REGION Network 8: Control the filling valve
         A     #Temp_IO_Status.HM_FillingValve;
         S     #Temp_IO_Status.HM_FillingValve1;
         S     #Temp_IO_Status.HM_FillingValve2;
   //
         AN    #Temp_IO_Status.HM_FillingValve;
         AN    #IN_Max_Level_Tank;
         R     #Temp_IO_Status.HM_FillingValve1;
         R     #Temp_IO_Status.HM_FillingValve2;
   //
         AN    #Temp_IO_Status.HM_FillingValve;
         AN    #Temp_IO_Status.HMFillingValves_Open;
         A     #Temp_IO_Status.V_FillingValve1;
         A     #Temp_IO_Status.V_FillingValve2;
         S     #Temp_IO_Status.HMFillingValves_Open;
   //
         A     #Temp_IO_Status.HMFillingValves_Open;
         L     S5T#3S;
         SP    #IN_Timer_Overlap_Valves;
   //
         AN    #Temp_IO_Status.HM_FillingValve;
         A     #Temp_IO_Status.V_FillingValve1;
         A     #Temp_IO_Status.V_FillingValve2;
         A     #Temp_IO_Status.HMFillingValves_Open;
         AN    #IN_Timer_Overlap_Valves;
         R     #Temp_IO_Status.HMFillingValves_Open;
   //
         AN    #Temp_IO_Status.HM_FillingValve;
         A     #Temp_IO_Status.HMFillingValves_Open;
         R     #Temp_IO_Status.HM_FillingValve1;
   //
         AN    #Temp_IO_Status.HM_FillingValve;
         AN    #Temp_IO_Status.HMFillingValves_Open;
         R     #Temp_IO_Status.HM_FillingValve2;
   //
         A     #Temp_IO_Status.HM_FillingValve1;
         L     S5T#2S;
         SF    #IN_Timer_Valve1;
   //
         A     #IN_Timer_Valve1;
         =     #Temp_IO_Status.V_FillingValve1;
   //
         A     #Temp_IO_Status.HM_FillingValve2;
         L     S5T#2S;
         SF    #IN_Timer_Valve2;
   //
         A     #IN_Timer_Valve2;
         =     #Temp_IO_Status.V_FillingValve2;
   //
         A     #Temp_IO_Status.V_FillingValve1;
         =     #OUT_FillingValve1;
   //
         A     #Temp_IO_Status.V_FillingValve2;
         =     #OUT_FillingValve2;
END_REGION

REGION Network 9
         AN    #Temp_IO_Status.V_FillingValve1;
   //    U     "E_FuellVent1_K1_geschl"
         AN    #Temp_IO_Status.HM_Valve2_closed;
         S     #Temp_IO_Status.HM_Valve1_closed;
   //
         AN    #Temp_IO_Status.V_FillingValve2;
   //    U     "E_FuellVent2_K1_geschl"
         AN    #Temp_IO_Status.HM_Valve1_closed;
         S     #Temp_IO_Status.HM_Valve2_closed;
   //
         A     #Temp_IO_Status.V_FillingValve1;
   //    U     "E_FuellVent1_K1_offen"
         R     #Temp_IO_Status.HM_Valve1_closed;
   //
         A     #Temp_IO_Status.V_FillingValve2;
   //    U     "E_FuellVent2_K1_offen"
         R     #Temp_IO_Status.HM_Valve1_closed;
   //
         A     #Temp_IO_Status.EnableComponentPump;
         AN    #IN_Max_Level_Tank;
         AN    #Temp_IO_Fault.FLT_Valve1_Max;
         S     #Temp_IO_Fault.FLT_Valve1_Max;
         S     #IO_FaultLevel_3;
   //-----
         A     #Temp_IO_Status.HM_Valve2_closed;
         AN    #IN_Max_Level_Tank;
         AN    #Temp_IO_Fault.FLT_Valve2_Max;
         S     #Temp_IO_Fault.FLT_Valve2_Max;
         S     #IO_FaultLevel_3;
   //-----
END_REGION

REGION Network 10: Save data
   Out:  NOP   0;
         CALL  BLKMOV
         ( SRCBLK  := #Temp_IO_Status,
           RET_VAL := #ERROR_CODE,
           DSTBLK  := #AnyPointer1
         );
   //-----
         CALL  BLKMOV
         ( SRCBLK  := #Temp_IO_Fault,
           RET_VAL := #ERROR_CODE,
           DSTBLK  := #AnyPointer2
         );
   //-----
END_REGION
END_FUNCTION

FUNCTION "Baustein_1" : Void   // FC3, SCL
{ S7_Optimized_Access := 'FALSE' }
VERSION : 0.1
   VAR_TEMP
      N : Int;
      Y : Int;
   END_VAR
BEGIN

   // Anzahl der Komponenten am Mischkopf und Zuweisung der Namen vom Tagesbehälter!
   // 
     "DB619_State_MPart".Recirculation[1].Lowpressure_Exist := 0;
     "DB619_State_MPart".Recirculation[2].Lowpressure_Exist := 0;

   FOR #N := 1 TO "DB790_PlantParameter".AmountMH DO
     // Statement section FOR

   "DB704_MH_Value".Mixinghead[#N].MH_Connection[1].Exist:=0;
   "DB704_MH_Value".Mixinghead[#N].MH_Connection[2].Exist:=0;
   "DB704_MH_Value".Mixinghead[#N].MH_Connection[3].Exist:=0;
   "DB704_MH_Value".Mixinghead[#N].MH_Connection[4].Exist:=0;
   "DB704_MH_Value".Mixinghead[#N].MH_Connection[5].Exist:=0;
   "DB704_MH_Value".Mixinghead[#N].MH_Connection[6].Exist:=0;

     IF "DB704_MH_Value".Mixinghead[#N].AmountComponent = 1 THEN
       "DB704_MH_Value".Mixinghead[#N].MH_Connection[1].Exist:=1;
     ELSIF "DB704_MH_Value".Mixinghead[#N].AmountComponent = 2 THEN
       "DB704_MH_Value".Mixinghead[#N].MH_Connection[1].Exist:=1; 
       "DB704_MH_Value".Mixinghead[#N].MH_Connection[2].Exist:=1;
     ELSIF "DB704_MH_Value".Mixinghead[#N].AmountComponent = 3 THEN
       "DB704_MH_Value".Mixinghead[#N].MH_Connection[1].Exist:=1;
       "DB704_MH_Value".Mixinghead[#N].MH_Connection[2].Exist:=1;
       "DB704_MH_Value".Mixinghead[#N].MH_Connection[3].Exist:=1;
     ELSIF "DB704_MH_Value".Mixinghead[#N].AmountComponent = 4 THEN
       "DB704_MH_Value".Mixinghead[#N].MH_Connection[1].Exist:=1; 
       "DB704_MH_Value".Mixinghead[#N].MH_Connection[2].Exist:=1;
       "DB704_MH_Value".Mixinghead[#N].MH_Connection[3].Exist:=1;
       "DB704_MH_Value".Mixinghead[#N].MH_Connection[4].Exist:=1;
     ELSIF "DB704_MH_Value".Mixinghead[#N].AmountComponent = 5 THEN
       "DB704_MH_Value".Mixinghead[#N].MH_Connection[1].Exist:=1;
       "DB704_MH_Value".Mixinghead[#N].MH_Connection[2].Exist:=1;
       "DB704_MH_Value".Mixinghead[#N].MH_Connection[3].Exist:=1;
       "DB704_MH_Value".Mixinghead[#N].MH_Connection[4].Exist:=1;
       "DB704_MH_Value".Mixinghead[#N].MH_Connection[5].Exist:=1;
     ELSIF "DB704_MH_Value".Mixinghead[#N].AmountComponent = 6 THEN
       "DB704_MH_Value".Mixinghead[#N].MH_Connection[1].Exist:=1;
       "DB704_MH_Value".Mixinghead[#N].MH_Connection[2].Exist:=1;
       "DB704_MH_Value".Mixinghead[#N].MH_Connection[3].Exist:=1;
       "DB704_MH_Value".Mixinghead[#N].MH_Connection[4].Exist:=1;
       "DB704_MH_Value".Mixinghead[#N].MH_Connection[5].Exist:=1;
       "DB704_MH_Value".Mixinghead[#N].MH_Connection[6].Exist:=1;
     END_IF;

   // Freigeben der Sollwert- Eingabe für den Durchfluß am Mischkopf
     "DB614_MH_State".MH_Status[#N].LP_Exist := 0;

     FOR #Y := 1 TO 6 DO
       "DB614_MH_State".MH_Connection[#N].Red_CircFlow_Exist[#Y] := 0;
       "DB614_MH_State".MH_Connection[#N].HP_CircFlow_Exist[#Y] := 0;
       "DB614_MH_State".MH_Connection[#N].LP_CircFlow_Exist[#Y] := 0;

       IF "DB704_MH_Value".Mixinghead[#N].MH_Connection[#Y].Exist = 1 THEN
         "DB614_MH_State".MH_Connection[#N].Red_CircFlow_Exist[#Y] := 1;
         "DB614_MH_State".MH_Connection[#N].HP_CircFlow_Exist[#Y] := 1;
         IF "DB704_MH_Value".Mixinghead[#N].WithLPCirculation = 1 THEN
           "DB614_MH_State".MH_Connection[#N].LP_CircFlow_Exist[#Y] := 1;
           "DB614_MH_State".MH_Status[#N].LP_Exist := 1;
         END_IF;
       END_IF;

   // Anzeige für kleine - Große Drehzahl
       "DB614_MH_State".MH_Connection[#N].HP_2Point_Flow_Exist[#Y]:= 0;
       "DB614_MH_State".MH_Connection[#N].Red_2Point_Flow_Exist[#Y]:= 0;
       "DB614_MH_State".MH_Connection[#N].LP_2Point_Flow_Exist[#Y]:= 0;

     IF "DB753_MeteringPump".Pump["DB704_MH_Value".Mixinghead[#N].MH_Connection[#Y].Pump_No].With_2Point THEN
       "DB614_MH_State".MH_Connection[#N].HP_2Point_Flow_Exist[#Y]:= "DB704_MH_Value".Mixinghead[#N].MH_Connection[#Y].Exist;
       "DB614_MH_State".MH_Connection[#N].Red_2Point_Flow_Exist[#Y]:= "DB704_MH_Value".Mixinghead[#N].MH_Connection[#Y].Exist;
       IF "DB704_MH_Value".Mixinghead[#N].WithLPCirculation = 1 THEN
         "DB614_MH_State".MH_Connection[#N].LP_2Point_Flow_Exist[#Y]:= "DB704_MH_Value".Mixinghead[#N].MH_Connection[#Y].Exist;
       END_IF;
     END_IF;

   // Anzeige für Düse/ Bypass- Ansteuerung
       "DB614_MH_State".MH_Connection[#N].Red_CircOverNozzle_Exist[#Y] := 0;
       "DB614_MH_State".MH_Connection[#N].HP_CircOverNozzle_Exist[#Y] := 0;
       "DB614_MH_State".MH_Connection[#N].LP_CircOverNozzle_Exist[#Y] := 0;

     IF "DB704_MH_Value".Mixinghead[#N].WithNozzleControl AND "DB704_MH_Value".Mixinghead[#N].MH_Connection[#Y].WithNozzle = 1 THEN
       "DB614_MH_State".MH_Connection[#N].Red_CircOverNozzle_Exist[#Y] := 1;
       "DB614_MH_State".MH_Connection[#N].HP_CircOverNozzle_Exist[#Y] := 1;
       IF "DB704_MH_Value".Mixinghead[#N].WithLPCirculation = 1 THEN
        "DB614_MH_State".MH_Connection[#N].LP_CircOverNozzle_Exist[#Y] := 1;
       END_IF;
     END_IF;

   // Anzeige der Eingaben für den schnellen Druckaufbau
     "DB614_MH_State".MH_Connection[#N].QPB_Exist[#Y] := 0;
     IF "DB614_MH_State".MH_Status[#N].QPB_Values_selected THEN
       "DB614_MH_State".MH_Connection[#N].QPB_Exist[#Y] := "DB704_MH_Value".Mixinghead[#N].MH_Connection[#Y].Exist;
     END_IF;

     END_FOR;

   // Taster für LowPressure anzeigen     
     IF "DB704_MH_Value".Mixinghead[#N].MachineNumber = 1 AND "DB614_MH_State".MH_Status[#N].LP_Exist THEN
       "DB619_State_MPart".Recirculation[1].Lowpressure_Exist := 1;
     ELSIF  "DB704_MH_Value".Mixinghead[#N].MachineNumber = 2 AND "DB614_MH_State".MH_Status[#N].LP_Exist THEN
       "DB619_State_MPart".Recirculation[2].Lowpressure_Exist := 1;
     END_IF;

   END_FOR;

   // Falls kein LowPressure existiert den Schalter ablöschen
     IF NOT "DB619_State_MPart".Recirculation[1].Lowpressure_Exist THEN
       "DB619_State_MPart".Recirculation[1].Switch_Lowpressure := 0;
     END_IF;
     IF NOT "DB619_State_MPart".Recirculation[2].Lowpressure_Exist THEN
       "DB619_State_MPart".Recirculation[2].Switch_Lowpressure := 0;
     END_IF;

   FOR #N := 1 TO "DB790_PlantParameter".AmountMH DO
     FOR #Y := 1 TO 6 DO
       // Anzeigen der Komponentennamen am Mischkopf
       "DB614_MH_State".MH_Connection[#N].Name[#Y] := "DB753_MeteringPump".Pump["DB704_MH_Value".Mixinghead[#N].MH_Connection[#Y].Pump_No].Name;

       // Anzeigen der Komponentenfarben am Mischkopf
       "DB614_MH_State".MH_Connection[#N].colour[#Y] := "DB613_Komponent_State".GroupStatus["DB704_MH_Value".Mixinghead[#N].MH_Connection[#Y].Pump_No].ColorTankFlow;

       // Begrenzen des minimal/maximal eingebbaren Durchflusses am Mischkopf
       "DB614_MH_State".MH_Connection[#N].MinFlow[#Y] := "DB613_Komponent_State".FlowPumpMin["DB704_MH_Value".Mixinghead[#N].MH_Connection[#Y].Pump_No];
       "DB614_MH_State".MH_Connection[#N].MaxFlow[#Y] := "DB613_Komponent_State".FlowPumpMax["DB704_MH_Value".Mixinghead[#N].MH_Connection[#Y].Pump_No];

       // Anzeige des aktuellen Durchflusses am Mischkopf
       "DB614_MH_State".MH_Connection[#N].ActFlow[#Y] := "DB608_PV_Metering".Metering["DB704_MH_Value".Mixinghead[#N].MH_Connection[#Y].Pump_No].Flow.PV_ActV.Value; 

     END_FOR;
   END_FOR;

   FOR #N := 1 TO "DB790_PlantParameter".AmountMH DO
   // Anzeige der Störungsinfo 
   "DB614_MH_State".MH_Status[#N].FaultExist := "DB614_MH_State".MH_CleaningPiston[#N].FaultExists;

   END_FOR;
END_FUNCTION

FUNCTION "FC4_Check_allocation" : Void   // FC4, SCL
{ S7_Optimized_Access := 'TRUE' }
VERSION : 0.1
// Function to check if selected program for delete is allocated
   VAR_INPUT
      Selected_tool : Int;   // Selected tool to delete
   END_VAR
   VAR_OUTPUT
      Delete_not_allowed : Bool;   // Delete not allowed. Tool is allocated
   END_VAR
   VAR_TEMP
      Ti_alloc_list : Int;
      TiLoop : Int;
      TiLoopMH : Int;
      Page : Int;
   END_VAR
BEGIN
   #Delete_not_allowed := FALSE;
   REGION automatic allocation list
       FOR #TiLoop := 1 TO "InterfaceVisu".AmountAlloactionAutomatic DO
           IF "DB940_Tool_alloc_automatic".Alloc_stationTool[#TiLoop] = #Selected_tool THEN
               #Delete_not_allowed := TRUE;
               "DB939_Tool_alloc_HMI".Tool_allocation_automatic := TRUE;
               "DB939_Tool_alloc_HMI".Select_hand_automatic_alloc := FALSE;
               "DB939_Tool_alloc_HMI".AllocList_page := (((#TiLoop-1) / 30) + 1);  // <-- Calculate page number
               "DB939_Tool_alloc_HMI".Selected_prog := #TiLoop - (((#TiLoop-1) / 30) * 30);  // Calculate place on actual list to set the focus
               RETURN;
           END_IF;
       END_FOR;
   END_REGION

   REGION manual allocation list MH
       FOR #TiLoopMH := 1 TO "DB790_PlantParameter".AmountMH DO
           IF "DB704_MH_Value".Mixinghead[#TiLoopMH].With99program THEN
               #Ti_alloc_list := 99;
           ELSE
               #Ti_alloc_list := 9;
           END_IF;

           FOR #TiLoop := 1 TO #Ti_alloc_list DO
               IF "DB941_Tool_alloc_manual_MH".MH[#TiLoopMH].Alloc_stationTool[#TiLoop] = #Selected_tool THEN
                   #Delete_not_allowed := TRUE;
                   "DB939_Tool_alloc_HMI".MH_No_selected := #TiLoopMH;
                   "DB939_Tool_alloc_HMI".Tool_allocation_manual := TRUE;
                   "DB939_Tool_alloc_HMI".Select_hand_automatic_alloc := TRUE;
                   "DB939_Tool_alloc_HMI".AllocList_page := (((#TiLoop-1) / 30) + 1);  // <-- Calculate page number
                   "DB939_Tool_alloc_HMI".Selected_prog := #TiLoop - (((#TiLoop-1) / 30) * 30);  // Calculate place on actual list to set the focus
                   RETURN;
               END_IF;
           END_FOR;
       END_FOR;
   END_REGION
END_FUNCTION

FUNCTION "FC5_Check_allocAutoMode" : Void   // FC5, SCL
{ S7_Optimized_Access := 'TRUE' }
VERSION : 0.1
   VAR_INPUT
      ToolcodeNo : Byte;   // Tool code number of the interface
   END_VAR
   VAR_OUTPUT
      ToolAlloc : Int;   // Allocation of the toolnumber to the allocation list
   END_VAR
BEGIN
   //---------------------------------------------------------------------------------------
   //Funktionsbeschreibung:
   //Diese Funktion wird verwendet, um zu übrprüfen, ob bei einer automatischen Werkzeugzuordnung über die Schnittstelle 
   //das entsprechende Werkzeug überhaupt gibt. Wenn es das Werkzeug nicht gibt, wird stattdessen die Werkzeug - Nummer 0 in die entsprechende Zuordnungsliste
   //geschrieben und eine Störmeldung an der Visualisierung angzeigt
   //----------------------------------------------------------------------------------------
   //

   REGION CheckToolNo
   // In diesem Abschnitt wird bei überprüft, ob es entsprechnedes Werkzeug vorhanden ist. Für die Überprüfung wird geschaut, ob im ersten Teilschuss
   // vom Werkzeug eine Mischkopfnummer (>0) vergeben ist
   // Ist das WErkzeug noch nicht erstellt wird eine entsprechende Fehlermeldung ausgegen
       IF "DB925_ShotData_1".Tool[#ToolcodeNo].Shot[1].MHNo > 0 THEN
           #ToolAlloc := BYTE_TO_INT(#ToolcodeNo);
       ELSE
           #ToolAlloc := 0;
           // Bilden der Fehlermeldung
       END_IF;
   END_REGION
END_FUNCTION

FUNCTION "FC011_OperationMode" : Void   // FC11, STL
TITLE = Operation mode
{ S7_Optimized_Access := 'FALSE' }
AUTHOR : KT242
FAMILY : RS_KK
NAME : BA
VERSION : 1.1
   VAR_INPUT
      IN_ContrVoltage : Bool;   // Signal control voltage on and emergency stop unlocked
      IN_Connection_OK : Bool;   // Communication to visualization is OK
      IN_SS_Manual : Bool;   // Input operation mode selector switch in manual mode
      IN_SS_Auto : Bool;   // Input operation mode selector switch in automatic mode
      IN_SS_Test : Bool;   // Input select testing flow of pumps by backflow valve
      IN_LampTest : Bool;   // Input to test lamp
      IN_Cycle_selected : Bool;   // Reciculation mode was activated by key
      IN_SS_CylinderService : Bool;   // Piston in service is selected by keyswitch
      IN_Hydraulic_OK : Bool;   // Feed back of hydraulic in operation
      IN_OperationMode_Timer : Timer;   // Timer to switch between operation modes
   END_VAR
   VAR_IN_OUT
      IO_Status : ANY;   // Save the operation mode
   END_VAR
   VAR_TEMP
      Temp_IO_Status : "UDT011_Operationmode";   // Local sate of operation mode to handle it iternal in the program block
      ERROR_CODE : Int;   // Error state of systemfunction "BLKMOV" Blockmove
      AnyPointer : ANY;   // Pointer to copy thr array "IO_Status" and "Temp_IO_Status"
   END_VAR
BEGIN

REGION Network 1: Saved data integration
   //-----
         LAR1;
         L;
         LAR2;
   //-----
         L     16#1002;  // Bytes
         T     W[AR1, P#0.0];
         L     W[AR2, P#2.0];  // Amount of bytes
         T     W[AR1, P#2.0];
         L     W[AR2, P#4.0];  // Block no,
         T     W[AR1, P#4.0];
         L     D[AR2, P#6.0];  // Startadress of datas
         T     D[AR1, P#6.0];
   //-----
         CALL  BLKMOV
         ( SRCBLK  := #AnyPointer,
           RET_VAL := #ERROR_CODE,
           DSTBLK  := #Temp_IO_Status
         );
   //-----
END_REGION

REGION Network 2: Operation mode selector-interpretation
   //-----
         A     #Temp_IO_Status.Controllvoltage;
         JC    Spg;
   //-----
         A     #IN_ContrVoltage;
         A     #IN_Connection_OK;
         L     S5T#1S;
         SD    #IN_OperationMode_Timer;
         A     #IN_OperationMode_Timer;
         =     #Temp_IO_Status.Controllvoltage;
         JU    BA;
   //-----
   Spg:  A     #IN_ContrVoltage;
         =     #Temp_IO_Status.Controllvoltage;
   //-----
         O(;
         AN    #IN_SS_Manual;
         A     #Temp_IO_Status.Manual;
         );
         O(;
         AN    #IN_SS_Auto;
         A     #Temp_IO_Status.Auto;
         );
         L     S5T#500MS;
         SE    #IN_OperationMode_Timer;
         A     #IN_OperationMode_Timer;
         JC    GOON;
   //-----
   BA:   A     #IN_SS_Manual;
         A     #Temp_IO_Status.Controllvoltage;
         =     #Temp_IO_Status.Manual;
   //-----
         A     #IN_SS_Auto;
         A     #Temp_IO_Status.Controllvoltage;
         =     #Temp_IO_Status.Auto;
   //-----
         A     #IN_SS_CylinderService;
         A     #Temp_IO_Status.Manual;
         AN    #IN_Cycle_selected;
         =     #Temp_IO_Status.Cylinderservice;
   //-----
         A     #IN_SS_Test;
         A     #Temp_IO_Status.Auto;
         =     #Temp_IO_Status.Test;
   //-----
   GOON: A     #IN_LampTest;
         A     #Temp_IO_Status.Controllvoltage;
         =     #Temp_IO_Status.Lamptest;
   //-----
         X     #Temp_IO_Status.SwitchOperation;
         X     #Temp_IO_Status.Operation;
         =     #Temp_IO_Status.Edge_OM_Change;
   //-----
         A     #Temp_IO_Status.SwitchOperation;
         =     #Temp_IO_Status.Operation;
   //-----
         O     #Temp_IO_Status.Manual;
         O     #Temp_IO_Status.Auto;
         =     #Temp_IO_Status.valid;
   //-----
         O     #Temp_IO_Status.Manual;
         O     #Temp_IO_Status.Auto;
         A     #IN_Hydraulic_OK;
         =     #Temp_IO_Status.Active;
   //-----
END_REGION

REGION Network 3: Save data
   //-----
         CALL  BLKMOV
         ( SRCBLK  := #Temp_IO_Status,
           RET_VAL := #ERROR_CODE,
           DSTBLK  := #AnyPointer
         );
   //-----
END_REGION
END_FUNCTION

FUNCTION "FC012_Circulation" : Void   // FC12, STL
TITLE = Circulation modes
{ S7_Optimized_Access := 'FALSE' }
AUTHOR : KT242
FAMILY : RS_KK
NAME : KRL
VERSION : 1.6
   VAR_INPUT
      IN_OperationMode_Manual : Bool;   // Foaming machine in manual mode
      IN_OperationMode_Auto : Bool;   // Foaming machine in automatic mode
      IN_OperationMode_active : Bool;   // Opearation mode is selected and hydraulic is active
      IN_Hydraulic_Switched_ON : Bool;   // Hydraulic was selected to switched on
      IN_Hydraulic_OK : Bool;   // Feed back of hydraulic in operation
      IN_LampTest : Bool;   // Input to test lamp
      IN_Cycle_running : Bool;   // Foaming cycle started
      IN_ShotPreparation_KK : Bool;   // Extarnel signal to fill component cylinder of a piston machine
      IN_Fault_Level_1 : Bool;   // Fault message of level 1 is active and was not acknowledged
      IN_Release_HP_Circ : Bool;   // General release of high pressure circulation
      IN_KK_in_PausingPos : Bool;   // Component cylinder in pausing position
      IN_Circulation_Timer : Timer;   // Timer for running and break during circulation at interval mode
      IN_Runtime_Manual : S5Time;   // Time value run-time of circulation at manual mode
      IN_Breaktime_Manual : S5Time;   // Time value break-time of circulation at manual mode
      IN_Runtime_Auto : S5Time;   // Time value run-time of circulation at automatic mode
      IN_Breaktime_Auto : S5Time;   // Time value braek-time of circulation at automatic mode
      IN_SWU_Release : "UDT001_DWord_1_32";   // Which switch over unit/mixing head is active at system
   END_VAR
   VAR_OUTPUT
      OU_MesIntervallTimeNOK : Bool;   // Message time value intervall mode not OK
   END_VAR
   VAR_IN_OUT
      IO_Status : ANY;   // Save status of circulation of the program
   END_VAR
   VAR_TEMP
      Temp_IO_Status : "UDT012_Recirculation";   // Internal status of circulation to work with at program block
      ERROR_CODE : Int;   // Error state of systemfunction "BLKMOV" Blockmove
      Anypointer : ANY;   // Pointer to copy thr array "IO_Status" and "Temp_IO_Status"
      Terminate_Circ : Bool;   // Termination-flag to stop circulaton during failure etc.
      Save_HighPressure : Bool;   // Intermidiate flag of HP-circulation to terminate cylinder machine
      Save_WeekendMode : Bool;   // Intermidiate flag of weekend-mode to terminate cylinder machine
      Save_ReducedCirc : Bool;   // Intermidiate flag of reduced-circulation to terminate cylinder machine
      Save_Interval : Bool;   // Intermidiate flag of run-time to terminate cylinder machine
      Save_Breaktime : Bool;   // Intermidiate flag of break-time to terminate cylinder machine
      Save_LowPressure : Bool;   // Intermidiate flag of low-pressure-circulation to terminate cylinder machine
      Save_CycleRuns : Bool;   // Intermidiate flag of active shot-cycle to terminate cylinder machine
      Programblock_No : Int;   // Flag to detect the memory area of the Bits "IN_SWU_Release"
      Address_ProgramBlock : DWord;   // and the start address within the program block
      Button_HP_local : DWord;   // Button at the mixinghead-panel to start high pressure-circulation
      Release_HP_local : DWord;   // Intermidiate flags of release of switch over units (from UDT to DWORD)
      Lamps_HP_local : DWord;   // Activation of high-pressure indicator at mixinghead-panel
      Temp_ReducedCirc_active : Bool;
      Temp_Intervall_active : Bool;
      Temp_LowPCirc_active : Bool;
      Temp_RunTimeManual : Time;
      Temp_BreakTimeManual : Time;
      Temp_RunTimeAuto : Time;
      Temp_BreakTimeAuto : Time;
      TempReleaseIntervall : Bool;
   END_VAR
BEGIN

REGION Network 1: Saved data integration
   // Änderungen:
   // -------------------------------------------------------------------------------
   // Befindet sich die Maschine im Kreislauf in der Pausenstellung und das 
   // Vorbereitungssignal vom Kolben kommt, sollte dieser ins Füllen gehen.
   // Dieses wurde das Einfügen des Eingangs "#IN_Schussvorbereitung_KK" im 
   // Netzwerk 4 Zeile 1 und das dadurch resultierende ablöschen der Pausenstellung 
   // erreicht.
   // 
   // Escher          10.08.2005
   // -------------------------------------------------------------------------------
   // Während der Pausenzeit im automatischen Intervall wurden die USE- Ventile nach 
   // Ablauf der Spülzeit umgeschaltet.
   // Geänderd durch einfügen der Zeile "UN    #Temp_IO_Status.Pausenzeit"
   // im Netzwerk 13 Zeile 9.
   // 
   // Grading         03.06.2004
   // -------------------------------------------------------------------------------
   // Bei einem angewählten ND- Kreislauf wurde die aktiv- Anzeige während der 
   // Pausenzeit nicht ausgeschaltet.
   // Geänderd durch einfügen der Zeile "UN    #Temp_IO_Status.Pausenzeit" 
   // im Netzwerk 14 Zeile 14.
   // 
   // v.d.Geest       27.10.2003
   // -------------------------------------------------------------------------------
   // Über das Bit "HD_ist_aktiv" und "Ist_aktiv" werden die Umschaltungen der USE- 
   // Ventile übernommen.
   // Nun kam es bei einem ausschalten des HD- Kreislaufes in den Stillstand der 
   // Maschine vor das genau für 1 SPS- Zyklus das Bit "ist_aktiv" noch gesetzt wurde 
   // aber "HD_ist_aktiv" nicht mehr. Hierdurch lief die Umschaltzeit und nicht die 
   // Abschaltzeit.
   // Also wird das Bit "Ist_aktiv" nun am Ende des Bausteins gesetzt.
   // 
   // v.d.Geest       11.04.2003
   // -------------------------------------------------------------------------------
   // Bei einer Störung der Gruppe 01 und einem angewähltem Kreislauf einer 
   // Pumpenmaschine wurden die Mischköpfe "durchgetaktet". Damit bei einer Störung 
   // keine Taktung mehr erfolgt wurde das Bit "Ist_aktiv" erstellt. Nur mit diesem 
   // Bit wird ein Takten der Mischköpfe vorgenommen.
   // Änderung des Bits "HD_angewaehlt" in "HD_ist_aktiv".
   // 
   // v.d.Geest       01.04.2003
   // -------------------------------------------------------------------------------
   //-----
         LAR1;
         L;
         LAR2;
   //-----
         L     W[AR2, P#0.0];  // Bytes
         T     W[AR1, P#0.0];
         L     W[AR2, P#2.0];  // Amount of bytes
         T     W[AR1, P#2.0];
         L     W[AR2, P#4.0];  // Block no,
         T     W[AR1, P#4.0];
         L     D[AR2, P#6.0];  // Startadress of datas
         T     D[AR1, P#6.0];
   //-----
         CALL  BLKMOV
         ( SRCBLK  := #Anypointer,
           RET_VAL := #ERROR_CODE,
           DSTBLK  := #Temp_IO_Status
         );
   //-----
END_REGION

REGION Network 2: Vorbelegung
   //-----
         A     #Temp_IO_Status.Intervall;
         =     #Save_Interval;
   //-----
         A     #Temp_IO_Status.Lowpressure;
         =     #Save_LowPressure;
   //-----
         A     #Temp_IO_Status.Reduced;
         =     #Save_ReducedCirc;
   //-----
         A     #Temp_IO_Status.Highpressure;
         =     #Save_HighPressure;
   //-----
         A     #Temp_IO_Status.Weekendswitching;
         =     #Save_WeekendMode;
   //-----
         A     #Temp_IO_Status.Pausetime;
         =     #Save_Breaktime;
   //-----
         A     #Temp_IO_Status.cycle_runs;
         =     #Save_CycleRuns;
   //-----
END_REGION

REGION Network 3: Circulation modes
   //-----
         AN    #IN_OperationMode_Auto;
         AN    #IN_OperationMode_Manual;
         ON    #IN_Hydraulic_OK;
         O     #IN_Fault_Level_1;
         AN    #Temp_IO_Status.Weekendswitching;
         =     #Terminate_Circ;
   //-----
         A     #IN_Cycle_running;
         =     #Temp_IO_Status.cycle_runs;
   //-----
         A     #Temp_IO_Status.HP_is_active;
         AN    #Terminate_Circ;
         =     #Temp_IO_Status.Highpressure;
   //-----
         A     #IN_OperationMode_Manual;
         A(;
         O     #Temp_IO_Status.Switch_Reduced;
         O     #Temp_IO_Status.Switch_Lowpressure;
         );
         A     #Temp_IO_Status.Switch_Intervall;
         AN    #Temp_IO_Status.Highpressure;
         A     #IN_Hydraulic_Switched_ON;
         =     #Temp_IO_Status.Weekendswitching;
   //-----
         A     #Temp_IO_Status.Switch_Reduced;
         AN    #Temp_IO_Status.Switch_Lowpressure;
         AN    #Temp_IO_Status.Highpressure;
         AN    #Terminate_Circ;
         =     #Temp_IO_Status.Reduced;
   //-----
         A     #Temp_IO_Status.Switch_Lowpressure;
         AN    #Temp_IO_Status.Highpressure;
         AN    #Terminate_Circ;
         =     #Temp_IO_Status.Lowpressure;
   //-----
END_REGION

REGION Network 4: Check time values intervall
   //-----
         CALL  T_CONV
         ( IN  := #IN_Runtime_Manual,
           OUT := #Temp_RunTimeManual
         );
   //-----
         CALL  T_CONV
         ( IN  := #IN_Breaktime_Manual,
           OUT := #Temp_BreakTimeManual
         );
   //-----
         CALL  T_CONV
         ( IN  := #IN_Runtime_Auto,
           OUT := #Temp_RunTimeAuto
         );
   //-----
         CALL  T_CONV
         ( IN  := #IN_Breaktime_Auto,
           OUT := #Temp_BreakTimeAuto
         );
   //-----
         A(;
         L     #Temp_RunTimeManual;
         L     0;
         >D;
         O     #IN_OperationMode_Auto;
         );
         A(;
         L     #Temp_BreakTimeManual;
         L     0;
         >D;
         O     #IN_OperationMode_Auto;
         );
         A(;
         L     #Temp_RunTimeAuto;
         L     0;
         >D;
         O     #IN_OperationMode_Manual;
         );
         A(;
         L     #Temp_BreakTimeAuto;
         L     0;
         >D;
         O     #IN_OperationMode_Manual;
         );
         =     #TempReleaseIntervall;
   //-----
         AN    #TempReleaseIntervall;
         =     #OU_MesIntervallTimeNOK;
   //-----
         O     #Temp_IO_Status.Reduced;
         O     #Temp_IO_Status.Lowpressure;
         A     #Temp_IO_Status.Switch_Intervall;
         A     #TempReleaseIntervall;
         =     #Temp_IO_Status.Intervall;
   //-----
END_REGION

REGION Network 5: The pouring machine is pausing time of the interval
   //-----
         O     #IN_ShotPreparation_KK;
         O     #Temp_IO_Status.cycle_runs;
         ON    #Temp_IO_Status.Intervall;
         R     #Temp_IO_Status.Pausetime;
         R     #Temp_IO_Status.RequestPausePos;
         R     #IN_Circulation_Timer;
         JC    TIME;
   //-----
         AN    #IN_Circulation_Timer;
         JC    BA;
   //-----
         AN    #Temp_IO_Status.Pausetime;
         AN    #IN_KK_in_PausingPos;
         =     #Temp_IO_Status.RequestPausePos;
         JC    Move;
   //-----
         AN    #Temp_IO_Status.Pausetime;
         A     #IN_KK_in_PausingPos;
         =     #Temp_IO_Status.Pausetime;
   //-----
   BA:   A     #IN_OperationMode_Auto;
         JC    AUTO;
   //-----
         L     #IN_Runtime_Manual;
         AN    #Temp_IO_Status.Pausetime;
         JC    TIME;
         L     #IN_Breaktime_Manual;
         JU    TIME;
   //-----
   AUTO: L     #IN_Runtime_Auto;
         AN    #Temp_IO_Status.Pausetime;
         JC    TIME;
         L     #IN_Breaktime_Auto;
   //-----
   TIME: A     #Temp_IO_Status.Intervall;
         AN    #Temp_IO_Status.cycle_runs;
         AN    #IN_Circulation_Timer;
         SD    #IN_Circulation_Timer;
   //-----
   Move: NOP   0;
END_REGION

REGION Network 6: Terminate circulation at piston machine
   //-----
         O(;
         X     #Temp_IO_Status.Highpressure;
         X     #Save_HighPressure;
         );
         O(;
         X     #Temp_IO_Status.Weekendswitching;
         X     #Save_WeekendMode;
         );
         O(;
         X     #Temp_IO_Status.Reduced;
         X     #Save_ReducedCirc;
         );
         O(;
         X     #Temp_IO_Status.Intervall;
         X     #Save_Interval;
         );
         O(;
         X     #Temp_IO_Status.Pausetime;
         X     #Save_Breaktime;
         AN    #Temp_IO_Status.Pausetime;
         );
         O(;
         X     #Temp_IO_Status.Lowpressure;
         X     #Save_LowPressure;
         );
         O     #IN_ShotPreparation_KK;
         AN    #Temp_IO_Status.cycle_runs;
         O(;
         X     #Temp_IO_Status.cycle_runs;
         X     #Save_CycleRuns;
         A     #Temp_IO_Status.cycle_runs;
         );
         =     #Temp_IO_Status.Break_KK;
   //-----
END_REGION

REGION Network 7
   //-----
         L;
         LAR1;
         L     W[AR1, P#0.0];
         T     #Programblock_No;
         L     D[AR1, P#2.0];
         T     #Address_ProgramBlock;
         LAR2;
         L;
         LAR1;
   //-----
         OPN   DB[ #Programblock_No];
         L     DBD[AR2, P#0.0];
         T     LD[AR1, P#0.0];
   //-----
   // Shift high pressure release to local DWord- area
   //-----
         L;
         LAR2;
         L;
         LAR1;
   //-----
         L     LD [ AR2 , P#16.0 ];
         T     LD[AR1, P#0.0];
   //-----
END_REGION

REGION Network 8: High pressure circulation of maximum 32 buttons
   //-----
         A(;
         L     #Temp_IO_Status.SWU_RC_HP;  // if SWU is deselected during
         L     #Release_HP_local;  // high pressure circulation
         AD;
         L     0;
         ==D;
         );
         A     #Temp_IO_Status.HP_is_active;
         ON    #IN_Release_HP_Circ;  // If their is no general release
         ON    #IN_OperationMode_active;
         O     #IN_Fault_Level_1;
         JC    DEL;  // than delete the state
   //-----
         L     #Temp_IO_Status.Status_RC_HP;
         JL    DEL;  // Jump list: Status_Circ. HP>3 Jump to DEL
         JU    FP1T;  // Button 0->1 : 1.time Status_Circ.-HP=0
         JU    FN1T;  // Button 1->0 : 1.time Status_Circ.-HP=1
         JU    FP2T;  // Button 0->1 : 2.time Status_Circ.-HP=2
         JU    FN2T;  // Button 1->0 : 2.time Status_Circ.-HP=3
   //-----
   DEL:  L     0;
         T     #Temp_IO_Status.SWU_RC_HP;
         T     #Temp_IO_Status.Status_RC_HP;
         JU    HDAN;
   //-----
END_REGION

REGION Network 9: Button 1.time pressed -> positive edge
   //-----
   FP1T: L     #Button_HP_local;  // Button 0->1
         L     #Release_HP_local;  // SWU release
         AD;
         T     #Temp_IO_Status.SWU_RC_HP;  // Activate SWU release for HP-Circulation
         L     0;
         >D;
         JCN   HDAN;
         L     1;
         T     #Temp_IO_Status.Status_RC_HP;
         JU    HDAN;
   //-----
END_REGION

REGION Network 10: Button 1.time pressed -> negative edge
   //-----
   FN1T: L     #Button_HP_local;  // Button 1->0
         L     0;
         ==D;
         JCN   HDAN;
         L     2;
         T     #Temp_IO_Status.Status_RC_HP;
         JU    HDAN;
   //-----
END_REGION

REGION Network 11: Button 2.time pressed -> positive edge
   //-----
   FP2T: L     #Button_HP_local;  //B utton 0->1
         L     #Temp_IO_Status.SWU_RC_HP;  // Button suits to SWU
         AD;
         L     0;
         >D;
         JCN   HDAN;
         L     3;
         T     #Temp_IO_Status.Status_RC_HP;
         JU    HDAN;
   //-----
END_REGION

REGION Network 12: Button 2.time pressed -> negative edge
   //-----
   FN2T: L     #Button_HP_local;  // Button 1->0
         L     #Temp_IO_Status.SWU_RC_HP;  // Button fits to SWU
         AD;
         L     0;
         ==D;
         JCN   HDAN;
         L     4;
         T     #Temp_IO_Status.Status_RC_HP;
         JU    HDAN;
   //-----
END_REGION

REGION Network 13: High pressure selected , Lamp activation
   //-----
   HDAN: L     #Temp_IO_Status.SWU_RC_HP;  // HP-Circulation is selected
         L     0;
         <>D;
         =     #Temp_IO_Status.HP_is_active;
   //-----
         A     #IN_LampTest;  // Test of indicator lights is selected
         L     16#0000_FFFF;
         JC    LAMP;
   //-----
         L     0;  // Lamps off
         A     #Temp_IO_Status.HP_is_active;
         AN    "Flag_01_000_Hertz";
         ON    #IN_Release_HP_Circ;
         JC    LAMP;
   //-----
         L     #Temp_IO_Status.SWU_RC_HP;  // Lamps as selected
         A     #Temp_IO_Status.HP_is_active;
         JC    LAMP;
   //-----
         L     #Release_HP_local;  // Lamps as released
   LAMP: NOP   0;
   //-----
         L;
         LAR2;
         TAK;
         T     LD [ AR2 , P#20.0 ];
   //-----
END_REGION

REGION Network 14: Output of active bits after selection of high pressure circ.
   //-----
         O     #Temp_IO_Status.Switch_Reduced;
         O     #Temp_IO_Status.Switch_Lowpressure;
         O     #Temp_IO_Status.HP_is_active;
         A     #IN_OperationMode_active;
         =     #Temp_IO_Status.Is_selected;
   //-----
         A     #Temp_IO_Status.Is_selected;
         AN    #IN_Fault_Level_1;
         AN    #Temp_IO_Status.Pausetime;
         =     #Temp_IO_Status.Is_active;
   //-----
END_REGION

REGION Network 15: Output of indication control at computer 1-> ON; 2-> Faulty; 3->Selected but not ON
   //-----
         A     #Temp_IO_Status.Reduced;
         A     #IN_OperationMode_active;
         AN    #Temp_IO_Status.Pausetime;
         AN    #IN_Cycle_running;
         AN    #IN_Fault_Level_1;
         =     #Temp_ReducedCirc_active;
   //-----
         A     #Temp_ReducedCirc_active;
         L     1;
         JC    Rtra;
   //-
         A     #IN_Fault_Level_1;
         L     2;
         JC    Rtra;
   //-
         AN    #Temp_ReducedCirc_active;
         A     #Temp_IO_Status.Switch_Reduced;
         L     3;
         JC    Rtra;
   //-
         L     0;
   Rtra: T     #Temp_IO_Status.State_Reduced;
   //-----
   //----- Intervall ----------------------
         A     #Temp_IO_Status.Intervall;
         AN    #IN_Cycle_running;
         =     #Temp_Intervall_active;
   //-----
         L     0;
         A     #Temp_Intervall_active;
         JCN   Ireq;
         L     1;
         JU    Itra;
   Ireq: A     #Temp_IO_Status.Switch_Intervall;
         AN    #Temp_Intervall_active;
         JCN   Itra;
         L     2;
   Itra: T     #Temp_IO_Status.State_Intervall;
   //-----
   //------ Low Pressure -------------------
         A     #Temp_IO_Status.Lowpressure;
         A     #IN_OperationMode_active;
         AN    #Temp_IO_Status.Pausetime;
         AN    #IN_Cycle_running;
         AN    #IN_Fault_Level_1;
         =     #Temp_LowPCirc_active;
   //-----
         A     #Temp_LowPCirc_active;
         L     1;
         JC    Ltra;
   //-
         A     #IN_Fault_Level_1;
         L     2;
         JC    Ltra;
   //-
         A     #Temp_IO_Status.Switch_Lowpressure;
         AN    #Temp_LowPCirc_active;
         L     2;
         JC    Ltra;
   //-
         L     0;
   Ltra: T     #Temp_IO_Status.State_Lowpressure;
   //-----
END_REGION

REGION Network 16: Save data
   //-----
         CALL  BLKMOV
         ( SRCBLK  := #Temp_IO_Status,
           RET_VAL := #ERROR_CODE,
           DSTBLK  := #Anypointer
         );
   //-----
END_REGION
END_FUNCTION

FUNCTION "FC14_TP_Shortcuts" : Void   // FC14, STL
{ S7_Optimized_Access := 'TRUE' }
VERSION : 0.1
BEGIN

REGION Network 1: Press Button vor 2 seconds will copy act page to set page
   // Any button pressed for 2 seconds
         O     "DB14_TP_Shortcuts".TP_Shortcuts.ButtonNo."1";
         O     "DB14_TP_Shortcuts".TP_Shortcuts.ButtonNo."2";
         O     "DB14_TP_Shortcuts".TP_Shortcuts.ButtonNo."3";
         O     "DB14_TP_Shortcuts".TP_Shortcuts.ButtonNo."4";
         O     "DB14_TP_Shortcuts".TP_Shortcuts.ButtonNo."5";
         O     "DB14_TP_Shortcuts".TP_Shortcuts.ButtonNo."6";
         O     "DB14_TP_Shortcuts".TP_Shortcuts.ButtonNo."7";

   // Block KM Setting pages
         AN(;
         O(;
         A(;
         L     "TP-Bereichszeiger".Picturenumber.Bildnummer;
         L     1000;  // 1000 Settings / 2000 Config
         >=I;
         );
         A(;
         L     "TP-Bereichszeiger".Picturenumber.Bildnummer;
         L     9000;  // Service pages = okay to store
         <I;
         );
         );
         O(;
         L     "TP-Bereichszeiger".Picturenumber.Bildnummer;
         L     5;  // Parameter mixing head
         ==I;
         );
         O(;
         L     "TP-Bereichszeiger".Picturenumber.Bildnummer;
         L     7;  // Parameter tanks
         ==I;
         );
         O(;
         L     "TP-Bereichszeiger".Picturenumber.Bildnummer;
         L     12;  // Parameter pumps
         ==I;
         );
         O(;
         L     "TP-Bereichszeiger".Picturenumber.Bildnummer;
         L     35;  // Parameter robot
         ==I;
         );

         );
         L     s5t#2s;
         SD    "T_Set_new_page_no";

         A     "T_Set_new_page_no";
         FP    "FP_new_page_no";
         JCN   end;

         A     "DB14_TP_Shortcuts".TP_Shortcuts.ButtonNo."1";
         JCN   B2;
         L     "TP-Bereichszeiger".Picturenumber.Bildnummer;
         L     "DB14_TP_Shortcuts".TP_Shortcuts.PageNo."1";
         ==I;
         L     0;
         JC    del1;
         L     "TP-Bereichszeiger".Picturenumber.Bildnummer;
   del1: T     "DB14_TP_Shortcuts".TP_Shortcuts.PageNo."1";

   B2:   A     "DB14_TP_Shortcuts".TP_Shortcuts.ButtonNo."2";
         JCN   B3;
         L     "TP-Bereichszeiger".Picturenumber.Bildnummer;
         L     "DB14_TP_Shortcuts".TP_Shortcuts.PageNo."2";
         ==I;
         L     0;
         JC    del2;
         L     "TP-Bereichszeiger".Picturenumber.Bildnummer;
   del2: T     "DB14_TP_Shortcuts".TP_Shortcuts.PageNo."2";

   B3:   A     "DB14_TP_Shortcuts".TP_Shortcuts.ButtonNo."3";
         JCN   B4;
         L     "TP-Bereichszeiger".Picturenumber.Bildnummer;
         L     "DB14_TP_Shortcuts".TP_Shortcuts.PageNo."3";
         ==I;
         L     0;
         JC    del3;
         L     "TP-Bereichszeiger".Picturenumber.Bildnummer;
   del3: T     "DB14_TP_Shortcuts".TP_Shortcuts.PageNo."3";

   B4:   A     "DB14_TP_Shortcuts".TP_Shortcuts.ButtonNo."4";
         JCN   B5;
         L     "TP-Bereichszeiger".Picturenumber.Bildnummer;
         L     "DB14_TP_Shortcuts".TP_Shortcuts.PageNo."4";
         ==I;
         L     0;
         JC    del4;
         L     "TP-Bereichszeiger".Picturenumber.Bildnummer;
   del4: T     "DB14_TP_Shortcuts".TP_Shortcuts.PageNo."4";

   B5:   A     "DB14_TP_Shortcuts".TP_Shortcuts.ButtonNo."5";
         JCN   B6;
         L     "TP-Bereichszeiger".Picturenumber.Bildnummer;
         L     "DB14_TP_Shortcuts".TP_Shortcuts.PageNo."5";
         ==I;
         L     0;
         JC    del5;
         L     "TP-Bereichszeiger".Picturenumber.Bildnummer;
   del5: T     "DB14_TP_Shortcuts".TP_Shortcuts.PageNo."5";

   B6:   A     "DB14_TP_Shortcuts".TP_Shortcuts.ButtonNo."6";
         JCN   B7;
         L     "TP-Bereichszeiger".Picturenumber.Bildnummer;
         L     "DB14_TP_Shortcuts".TP_Shortcuts.PageNo."6";
         ==I;
         L     0;
         JC    del6;
         L     "TP-Bereichszeiger".Picturenumber.Bildnummer;
   del6: T     "DB14_TP_Shortcuts".TP_Shortcuts.PageNo."6";

   B7:   A     "DB14_TP_Shortcuts".TP_Shortcuts.ButtonNo."7";
         JCN   B8;
         L     "TP-Bereichszeiger".Picturenumber.Bildnummer;
         L     "DB14_TP_Shortcuts".TP_Shortcuts.PageNo."7";
         ==I;
         L     0;
         JC    del7;
         L     "TP-Bereichszeiger".Picturenumber.Bildnummer;
   del7: T     "DB14_TP_Shortcuts".TP_Shortcuts.PageNo."7";

   B8:   NOP   0;

   end:  NOP   0;
END_REGION

REGION Network 2: Check if selected page is active

         L     "TP-Bereichszeiger".Picturenumber.Bildnummer;
         L     "DB14_TP_Shortcuts".TP_Shortcuts.PageNo."1";
         ==I;
         =     "DB14_TP_Shortcuts".TP_Shortcuts.Page_active."1";

         L     "TP-Bereichszeiger".Picturenumber.Bildnummer;
         L     "DB14_TP_Shortcuts".TP_Shortcuts.PageNo."2";
         ==I;
         =     "DB14_TP_Shortcuts".TP_Shortcuts.Page_active."2";

         L     "TP-Bereichszeiger".Picturenumber.Bildnummer;
         L     "DB14_TP_Shortcuts".TP_Shortcuts.PageNo."3";
         ==I;
         =     "DB14_TP_Shortcuts".TP_Shortcuts.Page_active."3";

         L     "TP-Bereichszeiger".Picturenumber.Bildnummer;
         L     "DB14_TP_Shortcuts".TP_Shortcuts.PageNo."4";
         ==I;
         =     "DB14_TP_Shortcuts".TP_Shortcuts.Page_active."4";

         L     "TP-Bereichszeiger".Picturenumber.Bildnummer;
         L     "DB14_TP_Shortcuts".TP_Shortcuts.PageNo."5";
         ==I;
         =     "DB14_TP_Shortcuts".TP_Shortcuts.Page_active."5";

         L     "TP-Bereichszeiger".Picturenumber.Bildnummer;
         L     "DB14_TP_Shortcuts".TP_Shortcuts.PageNo."6";
         ==I;
         =     "DB14_TP_Shortcuts".TP_Shortcuts.Page_active."6";

         L     "TP-Bereichszeiger".Picturenumber.Bildnummer;
         L     "DB14_TP_Shortcuts".TP_Shortcuts.PageNo."7";
         ==I;
         =     "DB14_TP_Shortcuts".TP_Shortcuts.Page_active."7";
END_REGION
END_FUNCTION

FUNCTION "FC021_MH_Hydraulic" : Void   // FC21, STL
TITLE = MH-Hydraulic
{ S7_Optimized_Access := 'FALSE' }
AUTHOR : KT242
FAMILY : RS_KK
NAME : MK_Hyd
VERSION : 1.1
   VAR_INPUT
      IN_MotorProtection : Bool;   // Input: Motorprotection hydraulic drive motor
      IN_Min_Level : Bool;   // Input: Minimum level of hydraulic oil was droped
      IN_C_OilCooling : Bool;   // Input: Temperature of oil exceed switchpoint oil-cooling valve on
      IN_C_Max : Bool;   // Input: Maximum temperature of hydraulic oil was exceeded->Warning-errormessage
      IN_F_Filter_FeedLine : Bool;   // Input: Pre flow high pressure filter is polluted
      IN_F_Filter_ReturnLine : Bool;   // Input: Back flow filter is polluted
      IN_OPMode_Automatic : Bool;   // Input: Foaming machine in automatic mode
      IN_OPMode_Manual : Bool;   // Input: Foaming machine in manual mode
      IN_PauseTime : Bool;   // Input: Foaming machine in pause time (Manual or Automatic)
      IN_Pos_of_Pause_ok : Bool;   // Input: Component pistons are in pause position
      IN_Fault_from_Extern : Bool;   // Input: External fault sswitch off hydraulic
      IN_P_lowerlimit : Bool;   // Input: Lower pressure limit hydraulic pressure reached
      IN_P_upperLimit : Bool;   // Input: Upper pressure limit hydraulic pressure not reached
      IN_Option2SetPoints : Bool;   // Option 2 setpoints for the hydraulic pressure used
      IN_PRequestCycle : Bool;   // Request pressure valve during foaming cycle
      IN_KK_Manager_active : Bool;   // Signal to use pistons to build up pressure
      IN_ShotStroke_by_Piston : Bool;   // Only during shot stroke of piston pressure valve is activated
      IN_Reset_fault_Fkt : Bool;   // Signal to acknowledge faults in functionblock
      IN_Temperatur_Timer : Timer;   // Timer duration of temperature warning after this temperature error
      IN_Filter_Timer : Timer;   // Timer delay fault high pressure-filter
      IN_Hydraulictimer : Timer;   // Timer to star up motors, pressure monitoring, and so on
      IN_Star_Delta_Timer : S5Time;   // Timevalue stat up hydraulic motor (star-delta starter)
      IN_Delay_FilterError : S5Time;   // Timevalue of delay filter error
      IN_P_BuildUpTime : S5Time;   // Timevalue monitoring pressure build up during switch on machine
      IN_P_OperationTime : S5Time;   // Timevalue monitoring pressure build up during normale operation machine
      IN_P_ClPistonTime : S5Time;   // Timevalue extension pressure build up request dof cleaning piston MH
      IN_SwitchOffTime : S5Time;
      IN_SwitchOFFTimer : Timer;
   END_VAR
   VAR_OUTPUT
      OUT_Hydraulic_active : Bool;   // Indicator hydraulic ready for operation
      OUT_PressureValve : Bool;   // Output pressure build up valve hydraulic
      OUT_Motor_MainsContactor : Bool;   // Output mains conactor hydraulic motor
      OUT_Motor_Star : Bool;   // Output of star contactor hydraulic motor
      OUT_Motor_Delta : Bool;   // Output of delta contactor hydraulic motor
      OUT_V_OilCooling : Bool;   // Output cooling valve hydraulic oil
   END_VAR
   VAR_IN_OUT
      IO_Status : ANY;   // Storage of operating status mixinghead hydraulic
      IO_Fault : ANY;
      IO_NewFault : Bool;
      IO_FaultLevel_1 : Bool;
      IO_FaultLevel_2 : Bool;
      IO_FaultLevel_3 : Bool;
   END_VAR
   VAR_TEMP
      Temp_IO_Status : "UDT021_Hydr_State";
      Temp_IO_Fault : "UDT1821_FLT_MH_Hydraulic";
      ERROR_CODE : Int;   // Error state of systemfunction "BLKMOV" Blockmove
      Anyzeiger1 : ANY;   // Pointer to copy thr array "IO_Status" and "Temp_IO_Status"
      Anyzeiger2 : ANY;   // Pointer to copy thr array "IO_Status" and "Temp_IO_Status"
      Temp_Motor_ON : S5Time;
      Temp_Motor_ON_ms : Time;
      Temp_Fault_Hyd : Bool;
      Temp_No_switch_OFF : Bool;
      Temp_Motor_ON_Auto : Bool;
      Temp_Switch_Motor_ON : Bool;
      Temp_DelayTimeZero : Bool;
   END_VAR
BEGIN

REGION Network 1: Saved data integration
   //-----
         LAR1;
         L;
         LAR2;
   //-----
         L     W[AR2, P#0.0];  // Bytes
         T     W[AR1, P#0.0];
         L     W[AR2, P#2.0];  // Amount of bytes
         T     W[AR1, P#2.0];
         L     W[AR2, P#4.0];  // Block no,
         T     W[AR1, P#4.0];
         L     D[AR2, P#6.0];  // Startadress of datas
         T     D[AR1, P#6.0];
   //-----
         CALL  BLKMOV
         ( SRCBLK  := #Anyzeiger1,
           RET_VAL := #ERROR_CODE,
           DSTBLK  := #Temp_IO_Status
         );
   //-----
         LAR1;
         L;
         LAR2;
   //-----
         L     W[AR2, P#0.0];  // Bytes
         T     W[AR1, P#0.0];
         L     W[AR2, P#2.0];  // Amount of bytes
         T     W[AR1, P#2.0];
         L     W[AR2, P#4.0];  // Block no,
         T     W[AR1, P#4.0];
         L     D[AR2, P#6.0];  // Startadress of datas
         T     D[AR1, P#6.0];
   //-----
         CALL  BLKMOV
         ( SRCBLK  := #Anyzeiger2,
           RET_VAL := #ERROR_CODE,
           DSTBLK  := #Temp_IO_Fault
         );
   //-----
END_REGION

